DATA_BLOCK "DB_SDC_TS_PARAMETER_6"   // DB3709
{ S7_Optimized_Access := 'FALSE' }
AUTHOR : FFM
FAMILY : SDC
NAME : SECT_DEF
VERSION : 1.0
   VAR
      HEADER : Struct   // Struktur für Datenheader // nicht verschieben
         DB_NR : Int := 3709;   // DB Nummer
         MIN_NR_SEK : Int := 501;   // Niedrigste SEK Nummer im DB
         MAX_NR_SEK : Int := 600;   // Höchste SEK Nummer im DB
         START_DAT : Int := 20;   // Startadresse der SEK im DB
         LAENGE_SEK_DATA : Int := 260;   // Länge SEK Data
         ANZ_PROFIL : Int := 10;   // Number of Profiles
         OFFEST_PROFIL : Int := 40;   // Offestadresse der Profilparameter im TS-Parameterdatensatz
         LAENGE_PROFIL_DATA : Int := 22;   // Länge SEK Data
         Res160 : Int := 0;   // Reserve
         Res : Int := 0;   // Reserve
      END_STRUCT;
      TS : Array[501..600] of "UDT_SDC_TS_PARAMETER";
   END_VAR
BEGIN
   TS[501].ALLG.SEK_NEXT_1 := 0;
   TS[501].ALLG.SEK_NEXT_2 := 0;
   TS[501].ALLG.Spare[4] := 16#00;
   TS[501].ALLG.Spare[5] := 16#00;
   TS[501].ALLG.POS.Start_1 := 1639750;
   TS[501].ALLG.POS.End_1 := 1646749;
   TS[501].ALLG.POS.Start_2 := 0;
   TS[501].ALLG.POS.End_2 := 0;
   TS[501].ALLG.POS.Actionpoint_1 := 0;
   TS[501].ALLG.POS.Actionpoint_2 := 0;
   TS[501].ALLG.FLAGS.DIST_VAL[0] := FALSE;
   TS[501].ALLG.FLAGS.DIST_VAL[1] := FALSE;
   TS[501].ALLG.FLAGS.DIST_VAL[2] := FALSE;
   TS[501].ALLG.FLAGS.DIST_VAL[3] := FALSE;
   TS[501].ALLG.FLAGS.DIST_VAL[4] := FALSE;
   TS[501].ALLG.FLAGS.DIST_VAL[5] := FALSE;
   TS[501].ALLG.FLAGS.DIST_VAL[6] := FALSE;
   TS[501].ALLG.FLAGS.DIST_VAL[7] := FALSE;
   TS[501].ALLG.FLAGS.DIST_VAL[8] := FALSE;
   TS[501].ALLG.FLAGS.DIST_VAL[9] := TRUE;
   TS[501].ALLG.FLAGS.DIST_VAL[10] := FALSE;
   TS[501].ALLG.FLAGS.DIST_VAL[11] := FALSE;
   TS[501].ALLG.FLAGS.DIST_VAL[12] := FALSE;
   TS[501].ALLG.FLAGS.DIST_VAL[13] := FALSE;
   TS[501].ALLG.FLAGS.DIST_VAL[14] := FALSE;
   TS[501].ALLG.FLAGS.DIST_VAL[15] := FALSE;
   TS[501].ALLG.FLAGS.one_profile := FALSE;
   TS[501].ALLG.FLAGS.BLIND := FALSE;
   TS[501].ALLG.FLAGS.NO_DIST_CONT := FALSE;
   TS[501].ALLG.FLAGS.SYNCH_AREA := FALSE;
   TS[501].ALLG.FLAGS.bit24 := FALSE;
   TS[501].ALLG.FLAGS.bit25 := FALSE;
   TS[501].ALLG.FLAGS.bit26 := FALSE;
   TS[501].ALLG.FLAGS.bit27 := FALSE;
   TS[501].ALLG.FLAGS.EN_HOIST := FALSE;
   TS[501].ALLG.FLAGS.D_RESET_AFTER := FALSE;
   TS[501].ALLG.FLAGS.D_PULK := FALSE;
   TS[501].ALLG.FLAGS.bit33 := FALSE;
   TS[501].ALLG.FLAGS.bit34 := FALSE;
   TS[501].ALLG.FLAGS.bit35 := FALSE;
   TS[501].ALLG.FLAGS.bit36 := FALSE;
   TS[501].ALLG.FLAGS.Deutronic_ON := FALSE;
   TS[501].ALLG.Stop_Position := 6500;
   TS[501].ALLG.Drive_speed_1 := 15000;
   TS[501].ALLG.Drive_speed_2 := 6000;
   TS[501].PROFIL[1].Hoist_Pos_start := 0;
   TS[501].PROFIL[1].Height := 3890;
   TS[501].PROFIL[1].Hoist_speed := 2000;
   TS[501].PROFIL[1].Hoist_offset_1 := 0;
   TS[501].PROFIL[1].Hoist_offset_2 := 0;
   TS[501].PROFIL[1].Hoist_offset_3 := 0;
   TS[501].PROFIL[1].Hoist_offset_4 := 0;
   TS[501].PROFIL[1].Hoist_Start_offset_1 := 0;
   TS[501].PROFIL[1].Hoist_Start_offset_2 := 0;
   TS[501].PROFIL[1].Hoist_Start_offset_3 := 0;
   TS[501].PROFIL[1].Hoist_Start_offset_4 := 0;
   TS[501].PROFIL[2].Hoist_Pos_start := 0;
   TS[501].PROFIL[2].Height := 3890;
   TS[501].PROFIL[2].Hoist_speed := 2000;
   TS[501].PROFIL[2].Hoist_offset_1 := 0;
   TS[501].PROFIL[2].Hoist_offset_2 := 0;
   TS[501].PROFIL[2].Hoist_offset_3 := 0;
   TS[501].PROFIL[2].Hoist_offset_4 := 0;
   TS[501].PROFIL[2].Hoist_Start_offset_1 := 0;
   TS[501].PROFIL[2].Hoist_Start_offset_2 := 0;
   TS[501].PROFIL[2].Hoist_Start_offset_3 := 0;
   TS[501].PROFIL[2].Hoist_Start_offset_4 := 0;
   TS[501].PROFIL[3].Hoist_Pos_start := 0;
   TS[501].PROFIL[3].Height := 3890;
   TS[501].PROFIL[3].Hoist_speed := 2000;
   TS[501].PROFIL[3].Hoist_offset_1 := 0;
   TS[501].PROFIL[3].Hoist_offset_2 := 0;
   TS[501].PROFIL[3].Hoist_offset_3 := 0;
   TS[501].PROFIL[3].Hoist_offset_4 := 0;
   TS[501].PROFIL[3].Hoist_Start_offset_1 := 0;
   TS[501].PROFIL[3].Hoist_Start_offset_2 := 0;
   TS[501].PROFIL[3].Hoist_Start_offset_3 := 0;
   TS[501].PROFIL[3].Hoist_Start_offset_4 := 0;
   TS[501].PROFIL[4].Hoist_Pos_start := 0;
   TS[501].PROFIL[4].Height := 3890;
   TS[501].PROFIL[4].Hoist_speed := 2000;
   TS[501].PROFIL[4].Hoist_offset_1 := 0;
   TS[501].PROFIL[4].Hoist_offset_2 := 0;
   TS[501].PROFIL[4].Hoist_offset_3 := 0;
   TS[501].PROFIL[4].Hoist_offset_4 := 0;
   TS[501].PROFIL[4].Hoist_Start_offset_1 := 0;
   TS[501].PROFIL[4].Hoist_Start_offset_2 := 0;
   TS[501].PROFIL[4].Hoist_Start_offset_3 := 0;
   TS[501].PROFIL[4].Hoist_Start_offset_4 := 0;
   TS[501].PROFIL[5].Hoist_Pos_start := 0;
   TS[501].PROFIL[5].Height := 3890;
   TS[501].PROFIL[5].Hoist_speed := 2000;
   TS[501].PROFIL[5].Hoist_offset_1 := 0;
   TS[501].PROFIL[5].Hoist_offset_2 := 0;
   TS[501].PROFIL[5].Hoist_offset_3 := 0;
   TS[501].PROFIL[5].Hoist_offset_4 := 0;
   TS[501].PROFIL[5].Hoist_Start_offset_1 := 0;
   TS[501].PROFIL[5].Hoist_Start_offset_2 := 0;
   TS[501].PROFIL[5].Hoist_Start_offset_3 := 0;
   TS[501].PROFIL[5].Hoist_Start_offset_4 := 0;
   TS[501].PROFIL[6].Hoist_Pos_start := 0;
   TS[501].PROFIL[6].Height := 3890;
   TS[501].PROFIL[6].Hoist_speed := 2000;
   TS[501].PROFIL[6].Hoist_offset_1 := 0;
   TS[501].PROFIL[6].Hoist_offset_2 := 0;
   TS[501].PROFIL[6].Hoist_offset_3 := 0;
   TS[501].PROFIL[6].Hoist_offset_4 := 0;
   TS[501].PROFIL[6].Hoist_Start_offset_1 := 0;
   TS[501].PROFIL[6].Hoist_Start_offset_2 := 0;
   TS[501].PROFIL[6].Hoist_Start_offset_3 := 0;
   TS[501].PROFIL[6].Hoist_Start_offset_4 := 0;
   TS[501].PROFIL[7].Hoist_Pos_start := 0;
   TS[501].PROFIL[7].Height := 3890;
   TS[501].PROFIL[7].Hoist_speed := 2000;
   TS[501].PROFIL[7].Hoist_offset_1 := 0;
   TS[501].PROFIL[7].Hoist_offset_2 := 0;
   TS[501].PROFIL[7].Hoist_offset_3 := 0;
   TS[501].PROFIL[7].Hoist_offset_4 := 0;
   TS[501].PROFIL[7].Hoist_Start_offset_1 := 0;
   TS[501].PROFIL[7].Hoist_Start_offset_2 := 0;
   TS[501].PROFIL[7].Hoist_Start_offset_3 := 0;
   TS[501].PROFIL[7].Hoist_Start_offset_4 := 0;
   TS[501].PROFIL[8].Hoist_Pos_start := 0;
   TS[501].PROFIL[8].Height := 3890;
   TS[501].PROFIL[8].Hoist_speed := 2000;
   TS[501].PROFIL[8].Hoist_offset_1 := 0;
   TS[501].PROFIL[8].Hoist_offset_2 := 0;
   TS[501].PROFIL[8].Hoist_offset_3 := 0;
   TS[501].PROFIL[8].Hoist_offset_4 := 0;
   TS[501].PROFIL[8].Hoist_Start_offset_1 := 0;
   TS[501].PROFIL[8].Hoist_Start_offset_2 := 0;
   TS[501].PROFIL[8].Hoist_Start_offset_3 := 0;
   TS[501].PROFIL[8].Hoist_Start_offset_4 := 0;
   TS[501].PROFIL[9].Hoist_Pos_start := 0;
   TS[501].PROFIL[9].Height := 3890;
   TS[501].PROFIL[9].Hoist_speed := 2000;
   TS[501].PROFIL[9].Hoist_offset_1 := 0;
   TS[501].PROFIL[9].Hoist_offset_2 := 0;
   TS[501].PROFIL[9].Hoist_offset_3 := 0;
   TS[501].PROFIL[9].Hoist_offset_4 := 0;
   TS[501].PROFIL[9].Hoist_Start_offset_1 := 0;
   TS[501].PROFIL[9].Hoist_Start_offset_2 := 0;
   TS[501].PROFIL[9].Hoist_Start_offset_3 := 0;
   TS[501].PROFIL[9].Hoist_Start_offset_4 := 0;
   TS[501].PROFIL[10].Hoist_Pos_start := 0;
   TS[501].PROFIL[10].Height := 3890;
   TS[501].PROFIL[10].Hoist_speed := 2000;
   TS[501].PROFIL[10].Hoist_offset_1 := 0;
   TS[501].PROFIL[10].Hoist_offset_2 := 0;
   TS[501].PROFIL[10].Hoist_offset_3 := 0;
   TS[501].PROFIL[10].Hoist_offset_4 := 0;
   TS[501].PROFIL[10].Hoist_Start_offset_1 := 0;
   TS[501].PROFIL[10].Hoist_Start_offset_2 := 0;
   TS[501].PROFIL[10].Hoist_Start_offset_3 := 0;
   TS[501].PROFIL[10].Hoist_Start_offset_4 := 0;
   TS[502].ALLG.SEK_NEXT_1 := 0;
   TS[502].ALLG.SEK_NEXT_2 := 0;
   TS[502].ALLG.Spare[4] := 16#00;
   TS[502].ALLG.Spare[5] := 16#00;
   TS[502].ALLG.POS.Start_1 := 1646750;
   TS[502].ALLG.POS.End_1 := 1653749;
   TS[502].ALLG.POS.Start_2 := 0;
   TS[502].ALLG.POS.End_2 := 0;
   TS[502].ALLG.POS.Actionpoint_1 := 0;
   TS[502].ALLG.POS.Actionpoint_2 := 0;
   TS[502].ALLG.FLAGS.DIST_VAL[0] := FALSE;
   TS[502].ALLG.FLAGS.DIST_VAL[1] := FALSE;
   TS[502].ALLG.FLAGS.DIST_VAL[2] := FALSE;
   TS[502].ALLG.FLAGS.DIST_VAL[3] := FALSE;
   TS[502].ALLG.FLAGS.DIST_VAL[4] := FALSE;
   TS[502].ALLG.FLAGS.DIST_VAL[5] := FALSE;
   TS[502].ALLG.FLAGS.DIST_VAL[6] := FALSE;
   TS[502].ALLG.FLAGS.DIST_VAL[7] := FALSE;
   TS[502].ALLG.FLAGS.DIST_VAL[8] := FALSE;
   TS[502].ALLG.FLAGS.DIST_VAL[9] := TRUE;
   TS[502].ALLG.FLAGS.DIST_VAL[10] := FALSE;
   TS[502].ALLG.FLAGS.DIST_VAL[11] := FALSE;
   TS[502].ALLG.FLAGS.DIST_VAL[12] := FALSE;
   TS[502].ALLG.FLAGS.DIST_VAL[13] := FALSE;
   TS[502].ALLG.FLAGS.DIST_VAL[14] := FALSE;
   TS[502].ALLG.FLAGS.DIST_VAL[15] := FALSE;
   TS[502].ALLG.FLAGS.one_profile := FALSE;
   TS[502].ALLG.FLAGS.BLIND := FALSE;
   TS[502].ALLG.FLAGS.NO_DIST_CONT := FALSE;
   TS[502].ALLG.FLAGS.SYNCH_AREA := FALSE;
   TS[502].ALLG.FLAGS.bit24 := FALSE;
   TS[502].ALLG.FLAGS.bit25 := FALSE;
   TS[502].ALLG.FLAGS.bit26 := FALSE;
   TS[502].ALLG.FLAGS.bit27 := FALSE;
   TS[502].ALLG.FLAGS.EN_HOIST := FALSE;
   TS[502].ALLG.FLAGS.D_RESET_AFTER := FALSE;
   TS[502].ALLG.FLAGS.D_PULK := FALSE;
   TS[502].ALLG.FLAGS.bit33 := FALSE;
   TS[502].ALLG.FLAGS.bit34 := FALSE;
   TS[502].ALLG.FLAGS.bit35 := FALSE;
   TS[502].ALLG.FLAGS.bit36 := FALSE;
   TS[502].ALLG.FLAGS.Deutronic_ON := FALSE;
   TS[502].ALLG.Stop_Position := 6400;
   TS[502].ALLG.Drive_speed_1 := 15000;
   TS[502].ALLG.Drive_speed_2 := 6000;
   // 15300 more start values not shown
END_DATA_BLOCK

DATA_BLOCK "DB_SDC_EMS_1"   // DB3714
{ S7_Optimized_Access := 'FALSE' }
VERSION : 0.1
   VAR
      HEADER : Struct
         DB_NR : Int := 3714;
         MIN_NR_EMS : Int := 1;
         MAX_NR_EMS : Int := 200;
         START_EMS : Int := 20;
         LAENGE_EMS : Int := 260;
         OFFSET_EMS_SEK_STAT : Int := 164;
         LAENGE_EMS_SEK_STAT : Int := 34;
         OFFSET_EMS_FKT : Int := 216;
         Res160 : Int := 0;
         Load : Bool := TRUE;
      END_STRUCT;
   END_VAR
BEGIN
END_DATA_BLOCK

DATA_BLOCK "DB_SDC_TS_IF_COMMAND"   // DB3716
{ S7_Optimized_Access := 'FALSE' }
AUTHOR : FFM
FAMILY : SDC
NAME : SECT_IF
VERSION : 0.1
   VAR
      HEADER : Struct   // Struktur für Datenheader // nicht verschieben
         DB_NR : Int := 3716;   // DB Nummer
         MIN_NR_SEK : Int := 1;   // Niedrigste SEK Nummer im DB
         MAX_NR_SEK : Int := 600;   // Höchste SEK Nummer im DB
         START_DAT : Int := 20;   // Startadresse der SEK im DB
         LAENGE_SEK_DATA : Int := 18;   // Länge SEK Data
         LAENGE_VAL_DATA : Int := 8;   // Länge Value Data
         LAENGE_BIT_DATA : Int := 6;   // Länge Bit Data
         LAENGE_FKT : Int := 4;   // Länge Funktion
         Res16 : Int;   // Reserve
         Res18 : Int;   // Reserve
      END_STRUCT;
      SEK : Array[1..600] of "UDT_SDC_EMS_TS_COM";   // Komando für Sektion
   END_VAR
BEGIN
END_DATA_BLOCK

DATA_BLOCK "DB_SDC_TS_IF_COMMAND_2"   // DB3717
{ S7_Optimized_Access := 'FALSE' }
AUTHOR : FFM
FAMILY : SDC
NAME : SECT_IF
VERSION : 0.1
   VAR
      HEADER : Struct   // Struktur für Datenheader // nicht verschieben
         DB_NR : Int := 3717;   // DB Nummer
         MIN_NR_SEK : Int := 601;   // Niedrigste SEK Nummer im DB
         MAX_NR_SEK : Int := 1000;   // Höchste SEK Nummer im DB
         START_DAT : Int := 20;   // Startadresse der SEK im DB
         LAENGE_SEK_DATA : Int := 18;   // Länge SEK Data
         LAENGE_VAL_DATA : Int := 8;   // Länge Value Data
         LAENGE_BIT_DATA : Int := 6;   // Länge Bit Data
         LAENGE_FKT : Int := 4;   // Länge Funktion
         Res16 : Int;   // Reserve
         Res18 : Int;   // Reserve
      END_STRUCT;
      SEK : Array[601..1000] of "UDT_SDC_EMS_TS_COM";   // Komando für Sektion
   END_VAR
BEGIN
END_DATA_BLOCK

DATA_BLOCK "DB_SDC_TS_IF_STATUS"   // DB3718
{ S7_Optimized_Access := 'FALSE' }
AUTHOR : FFM
FAMILY : SDC
NAME : SECT_IF
VERSION : 1.0
   VAR
      HEADER : Struct
         DB_NR : Int := 3718;
         MIN_NR_SEK : Int := 1;
         MAX_NR_SEK : Int := 600;
         START_DAT : Int := 20;
         LAENGE_SEK_DATA : Int := 34;
         LAENGE_VAL_DATA : Int := 18;
         LAENGE_BIT_DATA : Int := 8;
         LAENGE_SERIES : Int := 4;
         LAENGE_FKT : Int := 4;
         Res18 : Int := 0;
      END_STRUCT;
      SEK : Array[1..600] of "UDT_SDC_EMS_TS_STAT";
   END_VAR
BEGIN
   SEK[1].VAL.EMS_ID := 1;
   SEK[1].VAL.PROFIL := 1;
   SEK[1].VAL.DRIVE_POS := 581346;
   SEK[1].VAL.HOIST_POS := 4151;
   SEK[1].VAL.ERROR := 504;
   SEK[1].VAL.DRIVE_POS_PERC := 0;
   SEK[1].VAL.SEK := 1;
   SEK[1].BIT.PRESENT := TRUE;
   SEK[1].BIT.ERROR := TRUE;
   SEK[1].BIT.MAN_IR := TRUE;
   SEK[1].BIT.MORE_EMS_PRESENT := FALSE;
   SEK[1].BIT.ER_COMMAND := FALSE;
   SEK[1].BIT.W_DIST := FALSE;
   SEK[1].BIT.Spare_0_6 := FALSE;
   SEK[1].BIT.MESS_ACT := FALSE;
   SEK[1].BIT.D_MOVING := FALSE;
   SEK[1].BIT.D_NOT_MOVING := TRUE;
   SEK[1].BIT.H_MOVING := FALSE;
   SEK[1].BIT.H_NOT_MOVING := TRUE;
   SEK[1].BIT.X_MOVING := FALSE;
   SEK[1].BIT.X_NOT_MOVING := TRUE;
   SEK[1].BIT.D_IN_POS := FALSE;
   SEK[1].BIT.Spare_2_1 := FALSE;
   SEK[1].BIT.D_BEFOR_POS := FALSE;
   SEK[1].BIT.D_AFTER_POS := TRUE;
   SEK[1].BIT.D_GR_AP1 := TRUE;
   SEK[1].BIT.D_SM_AP1 := FALSE;
   SEK[1].BIT.D_GR_AP2 := TRUE;
   SEK[1].BIT.D_SM_AP2 := FALSE;
   SEK[1].BIT.H_IN_POS := TRUE;
   SEK[1].BIT.H_IN_TOPPOS := TRUE;
   SEK[1].BIT.H_IN_POS1 := FALSE;
   SEK[1].BIT.H_IN_POS2 := FALSE;
   SEK[1].BIT.H_IN_POS3 := FALSE;
   SEK[1].BIT.H_IN_POS4 := FALSE;
   SEK[1].BIT.H_GR_POS := FALSE;
   SEK[1].BIT.H_SM_POS := FALSE;
   SEK[1].BIT.H_GR_POS1 := FALSE;
   SEK[1].BIT.H_SM_POS1 := FALSE;
   SEK[1].BIT.H_GR_POS2 := FALSE;
   SEK[1].BIT.H_SM_POS2 := FALSE;
   SEK[1].BIT.H_GR_POS3 := FALSE;
   SEK[1].BIT.H_SM_POS3 := FALSE;
   SEK[1].BIT.H_GR_POS4 := FALSE;
   SEK[1].BIT.H_SM_POS4 := FALSE;
   SEK[1].BIT.H_BOTTOM_POS := FALSE;
   SEK[1].BIT.H_DISABLED := TRUE;
   SEK[1].BIT.H_CLEAR := FALSE;
   SEK[1].BIT.D_MOVING_FWD := FALSE;
   SEK[1].BIT.D_MOVING_RWD := FALSE;
   SEK[1].BIT.D_RESET_AFTER := FALSE;
   SEK[1].BIT.D_PULK := FALSE;
   SEK[1].BIT.D_NO_POS := FALSE;
   SEK[1].SORTE[1] := 'L';
   SEK[1].SORTE[2] := 'E';
   SEK[1].SORTE[3] := 'E';
   SEK[1].SORTE[4] := 'R';
   SEK[1].FKT.EMS_TO_REPAIR_1 := FALSE;
   SEK[1].FKT.EMS_TO_REPAIR_2 := FALSE;
   SEK[1].FKT.EMERG_HOIST := FALSE;
   SEK[1].FKT.Reserve_03 := FALSE;
   SEK[1].FKT.EMERG_DRIVE_FC := FALSE;
   SEK[1].FKT.Reserve_05 := FALSE;
   SEK[1].FKT.LAMP_TEST := FALSE;
   SEK[1].FKT.VAC_CLEAN := FALSE;
   SEK[1].FKT.PE_TEST := FALSE;
   SEK[1].FKT.KOHLE_TEST := FALSE;
   SEK[1].FKT.KOM_TEST := FALSE;
   SEK[1].FKT.Reserve_11 := FALSE;
   SEK[1].FKT.Reserve_12 := FALSE;
   SEK[1].FKT.Reserve_13 := FALSE;
   SEK[1].FKT.Reserve_14 := FALSE;
   SEK[1].FKT.Reserve_15 := FALSE;
   SEK[1].SPARE := 16#0000;
   SEK[2].VAL.EMS_ID := 0;
   SEK[2].VAL.PROFIL := 0;
   SEK[2].VAL.DRIVE_POS := 0;
   SEK[2].VAL.HOIST_POS := 0;
   SEK[2].VAL.ERROR := 0;
   SEK[2].VAL.DRIVE_POS_PERC := 0;
   SEK[2].VAL.SEK := 0;
   SEK[2].BIT.PRESENT := FALSE;
   SEK[2].BIT.ERROR := FALSE;
   SEK[2].BIT.MAN_IR := FALSE;
   SEK[2].BIT.MORE_EMS_PRESENT := FALSE;
   SEK[2].BIT.ER_COMMAND := FALSE;
   SEK[2].BIT.W_DIST := FALSE;
   SEK[2].BIT.Spare_0_6 := FALSE;
   SEK[2].BIT.MESS_ACT := FALSE;
   SEK[2].BIT.D_MOVING := FALSE;
   SEK[2].BIT.D_NOT_MOVING := FALSE;
   SEK[2].BIT.H_MOVING := FALSE;
   SEK[2].BIT.H_NOT_MOVING := FALSE;
   SEK[2].BIT.X_MOVING := FALSE;
   SEK[2].BIT.X_NOT_MOVING := FALSE;
   SEK[2].BIT.D_IN_POS := FALSE;
   SEK[2].BIT.Spare_2_1 := FALSE;
   SEK[2].BIT.D_BEFOR_POS := FALSE;
   SEK[2].BIT.D_AFTER_POS := FALSE;
   SEK[2].BIT.D_GR_AP1 := FALSE;
   SEK[2].BIT.D_SM_AP1 := FALSE;
   SEK[2].BIT.D_GR_AP2 := FALSE;
   SEK[2].BIT.D_SM_AP2 := FALSE;
   SEK[2].BIT.H_IN_POS := FALSE;
   SEK[2].BIT.H_IN_TOPPOS := FALSE;
   SEK[2].BIT.H_IN_POS1 := FALSE;
   SEK[2].BIT.H_IN_POS2 := FALSE;
   SEK[2].BIT.H_IN_POS3 := FALSE;
   SEK[2].BIT.H_IN_POS4 := FALSE;
   SEK[2].BIT.H_GR_POS := FALSE;
   SEK[2].BIT.H_SM_POS := FALSE;
   SEK[2].BIT.H_GR_POS1 := FALSE;
   SEK[2].BIT.H_SM_POS1 := FALSE;
   SEK[2].BIT.H_GR_POS2 := FALSE;
   SEK[2].BIT.H_SM_POS2 := FALSE;
   SEK[2].BIT.H_GR_POS3 := FALSE;
   SEK[2].BIT.H_SM_POS3 := FALSE;
   SEK[2].BIT.H_GR_POS4 := FALSE;
   SEK[2].BIT.H_SM_POS4 := FALSE;
   SEK[2].BIT.H_BOTTOM_POS := FALSE;
   SEK[2].BIT.H_DISABLED := FALSE;
   SEK[2].BIT.H_CLEAR := FALSE;
   SEK[2].BIT.D_MOVING_FWD := FALSE;
   SEK[2].BIT.D_MOVING_RWD := FALSE;
   SEK[2].BIT.D_RESET_AFTER := FALSE;
   SEK[2].BIT.D_PULK := FALSE;
   SEK[2].BIT.D_NO_POS := TRUE;
   SEK[2].SORTE[1] := ' ';
   SEK[2].SORTE[2] := ' ';
   SEK[2].SORTE[3] := ' ';
   SEK[2].SORTE[4] := ' ';
   SEK[2].FKT.EMS_TO_REPAIR_1 := FALSE;
   SEK[2].FKT.EMS_TO_REPAIR_2 := FALSE;
   SEK[2].FKT.EMERG_HOIST := FALSE;
   SEK[2].FKT.Reserve_03 := FALSE;
   SEK[2].FKT.EMERG_DRIVE_FC := FALSE;
   SEK[2].FKT.Reserve_05 := FALSE;
   SEK[2].FKT.LAMP_TEST := FALSE;
   SEK[2].FKT.VAC_CLEAN := FALSE;
   SEK[2].FKT.PE_TEST := FALSE;
   SEK[2].FKT.KOHLE_TEST := FALSE;
   SEK[2].FKT.KOM_TEST := FALSE;
   SEK[2].FKT.Reserve_11 := FALSE;
   SEK[2].FKT.Reserve_12 := FALSE;
   SEK[2].FKT.Reserve_13 := FALSE;
   SEK[2].FKT.Reserve_14 := FALSE;
   SEK[2].FKT.Reserve_15 := FALSE;
   SEK[2].SPARE := 16#0000;
   SEK[3].VAL.EMS_ID := 0;
   SEK[3].VAL.PROFIL := 0;
   SEK[3].VAL.DRIVE_POS := 0;
   SEK[3].VAL.HOIST_POS := 0;
   SEK[3].VAL.ERROR := 0;
   SEK[3].VAL.DRIVE_POS_PERC := 0;
   SEK[3].VAL.SEK := 0;
   SEK[3].BIT.PRESENT := FALSE;
   SEK[3].BIT.ERROR := FALSE;
   SEK[3].BIT.MAN_IR := FALSE;
   SEK[3].BIT.MORE_EMS_PRESENT := FALSE;
   SEK[3].BIT.ER_COMMAND := FALSE;
   SEK[3].BIT.W_DIST := FALSE;
   SEK[3].BIT.Spare_0_6 := FALSE;
   SEK[3].BIT.MESS_ACT := FALSE;
   SEK[3].BIT.D_MOVING := FALSE;
   SEK[3].BIT.D_NOT_MOVING := FALSE;
   SEK[3].BIT.H_MOVING := FALSE;
   SEK[3].BIT.H_NOT_MOVING := FALSE;
   SEK[3].BIT.X_MOVING := FALSE;
   SEK[3].BIT.X_NOT_MOVING := FALSE;
   SEK[3].BIT.D_IN_POS := FALSE;
   SEK[3].BIT.Spare_2_1 := FALSE;
   SEK[3].BIT.D_BEFOR_POS := FALSE;
   SEK[3].BIT.D_AFTER_POS := FALSE;
   SEK[3].BIT.D_GR_AP1 := FALSE;
   SEK[3].BIT.D_SM_AP1 := FALSE;
   SEK[3].BIT.D_GR_AP2 := FALSE;
   SEK[3].BIT.D_SM_AP2 := FALSE;
   SEK[3].BIT.H_IN_POS := FALSE;
   SEK[3].BIT.H_IN_TOPPOS := FALSE;
   SEK[3].BIT.H_IN_POS1 := FALSE;
   SEK[3].BIT.H_IN_POS2 := FALSE;
   SEK[3].BIT.H_IN_POS3 := FALSE;
   SEK[3].BIT.H_IN_POS4 := FALSE;
   SEK[3].BIT.H_GR_POS := FALSE;
   SEK[3].BIT.H_SM_POS := FALSE;
   SEK[3].BIT.H_GR_POS1 := FALSE;
   SEK[3].BIT.H_SM_POS1 := FALSE;
   SEK[3].BIT.H_GR_POS2 := FALSE;
   SEK[3].BIT.H_SM_POS2 := FALSE;
   SEK[3].BIT.H_GR_POS3 := FALSE;
   SEK[3].BIT.H_SM_POS3 := FALSE;
   SEK[3].BIT.H_GR_POS4 := FALSE;
   SEK[3].BIT.H_SM_POS4 := FALSE;
   SEK[3].BIT.H_BOTTOM_POS := FALSE;
   SEK[3].BIT.H_DISABLED := FALSE;
   SEK[3].BIT.H_CLEAR := FALSE;
   SEK[3].BIT.D_MOVING_FWD := FALSE;
   SEK[3].BIT.D_MOVING_RWD := FALSE;
   SEK[3].BIT.D_RESET_AFTER := FALSE;
   SEK[3].BIT.D_PULK := FALSE;
   // 44200 more start values not shown
END_DATA_BLOCK

DATA_BLOCK "DB_SDC_TS_IF_STATUS_2"   // DB3719
{ S7_Optimized_Access := 'FALSE' }
AUTHOR : FFM
FAMILY : SDC
NAME : SECT_IF
VERSION : 1.0
   VAR
      HEADER : Struct   // Struktur für Datenheader // nicht verschieben
         DB_NR : Int := 3719;   // DB Nummer
         MIN_NR_SEK : Int := 601;   // Niedrigste SEK Nummer im DB
         MAX_NR_SEK : Int := 1000;   // Höchste SEK Nummer im DB
         START_DAT : Int := 20;   // Startadresse der SEK im DB
         LAENGE_SEK_DATA : Int := 34;   // Länge SEK Data
         LAENGE_VAL_DATA : Int := 18;   // Länge Value Data
         LAENGE_BIT_DATA : Int := 8;   // Länge Bit Data
         LAENGE_SERIES : Int := 4;   // Länge SERIES
         LAENGE_FKT : Int := 4;   // Länge Funktion
         Res18 : Int := 0;   // Reserve
      END_STRUCT;
      SEK : Array[601..1000] of "UDT_SDC_EMS_TS_STAT";   // Status of section
   END_VAR
BEGIN
   SEK[601].VAL.EMS_ID := 0;
   SEK[601].VAL.PROFIL := 0;
   SEK[601].VAL.DRIVE_POS := 0;
   SEK[601].VAL.HOIST_POS := 0;
   SEK[601].VAL.ERROR := 0;
   SEK[601].VAL.DRIVE_POS_PERC := 0;
   SEK[601].VAL.SEK := 0;
   SEK[601].BIT.PRESENT := FALSE;
   SEK[601].BIT.ERROR := FALSE;
   SEK[601].BIT.MAN_IR := FALSE;
   SEK[601].BIT.MORE_EMS_PRESENT := FALSE;
   SEK[601].BIT.ER_COMMAND := FALSE;
   SEK[601].BIT.W_DIST := FALSE;
   SEK[601].BIT.Spare_0_6 := FALSE;
   SEK[601].BIT.MESS_ACT := FALSE;
   SEK[601].BIT.D_MOVING := FALSE;
   SEK[601].BIT.D_NOT_MOVING := FALSE;
   SEK[601].BIT.H_MOVING := FALSE;
   SEK[601].BIT.H_NOT_MOVING := FALSE;
   SEK[601].BIT.X_MOVING := FALSE;
   SEK[601].BIT.X_NOT_MOVING := FALSE;
   SEK[601].BIT.D_IN_POS := FALSE;
   SEK[601].BIT.Spare_2_1 := FALSE;
   SEK[601].BIT.D_BEFOR_POS := FALSE;
   SEK[601].BIT.D_AFTER_POS := FALSE;
   SEK[601].BIT.D_GR_AP1 := FALSE;
   SEK[601].BIT.D_SM_AP1 := FALSE;
   SEK[601].BIT.D_GR_AP2 := FALSE;
   SEK[601].BIT.D_SM_AP2 := FALSE;
   SEK[601].BIT.H_IN_POS := FALSE;
   SEK[601].BIT.H_IN_TOPPOS := FALSE;
   SEK[601].BIT.H_IN_POS1 := FALSE;
   SEK[601].BIT.H_IN_POS2 := FALSE;
   SEK[601].BIT.H_IN_POS3 := FALSE;
   SEK[601].BIT.H_IN_POS4 := FALSE;
   SEK[601].BIT.H_GR_POS := FALSE;
   SEK[601].BIT.H_SM_POS := FALSE;
   SEK[601].BIT.H_GR_POS1 := FALSE;
   SEK[601].BIT.H_SM_POS1 := FALSE;
   SEK[601].BIT.H_GR_POS2 := FALSE;
   SEK[601].BIT.H_SM_POS2 := FALSE;
   SEK[601].BIT.H_GR_POS3 := FALSE;
   SEK[601].BIT.H_SM_POS3 := FALSE;
   SEK[601].BIT.H_GR_POS4 := FALSE;
   SEK[601].BIT.H_SM_POS4 := FALSE;
   SEK[601].BIT.H_BOTTOM_POS := FALSE;
   SEK[601].BIT.H_DISABLED := FALSE;
   SEK[601].BIT.H_CLEAR := FALSE;
   SEK[601].BIT.D_MOVING_FWD := FALSE;
   SEK[601].BIT.D_MOVING_RWD := FALSE;
   SEK[601].BIT.D_RESET_AFTER := FALSE;
   SEK[601].BIT.D_PULK := FALSE;
   SEK[601].BIT.D_NO_POS := FALSE;
   SEK[601].SORTE[1] := ' ';
   SEK[601].SORTE[2] := ' ';
   SEK[601].SORTE[3] := ' ';
   SEK[601].SORTE[4] := ' ';
   SEK[601].FKT.EMS_TO_REPAIR_1 := FALSE;
   SEK[601].FKT.EMS_TO_REPAIR_2 := FALSE;
   SEK[601].FKT.EMERG_HOIST := FALSE;
   SEK[601].FKT.Reserve_03 := FALSE;
   SEK[601].FKT.EMERG_DRIVE_FC := FALSE;
   SEK[601].FKT.Reserve_05 := FALSE;
   SEK[601].FKT.LAMP_TEST := FALSE;
   SEK[601].FKT.VAC_CLEAN := FALSE;
   SEK[601].FKT.PE_TEST := FALSE;
   SEK[601].FKT.KOHLE_TEST := FALSE;
   SEK[601].FKT.KOM_TEST := FALSE;
   SEK[601].FKT.Reserve_11 := FALSE;
   SEK[601].FKT.Reserve_12 := FALSE;
   SEK[601].FKT.Reserve_13 := FALSE;
   SEK[601].FKT.Reserve_14 := FALSE;
   SEK[601].FKT.Reserve_15 := FALSE;
   SEK[601].SPARE := 16#0000;
   SEK[602].VAL.EMS_ID := 0;
   SEK[602].VAL.PROFIL := 0;
   SEK[602].VAL.DRIVE_POS := 0;
   SEK[602].VAL.HOIST_POS := 0;
   SEK[602].VAL.ERROR := 0;
   SEK[602].VAL.DRIVE_POS_PERC := 0;
   SEK[602].VAL.SEK := 0;
   SEK[602].BIT.PRESENT := FALSE;
   SEK[602].BIT.ERROR := FALSE;
   SEK[602].BIT.MAN_IR := FALSE;
   SEK[602].BIT.MORE_EMS_PRESENT := FALSE;
   SEK[602].BIT.ER_COMMAND := FALSE;
   SEK[602].BIT.W_DIST := FALSE;
   SEK[602].BIT.Spare_0_6 := FALSE;
   SEK[602].BIT.MESS_ACT := FALSE;
   SEK[602].BIT.D_MOVING := FALSE;
   SEK[602].BIT.D_NOT_MOVING := FALSE;
   SEK[602].BIT.H_MOVING := FALSE;
   SEK[602].BIT.H_NOT_MOVING := FALSE;
   SEK[602].BIT.X_MOVING := FALSE;
   SEK[602].BIT.X_NOT_MOVING := FALSE;
   SEK[602].BIT.D_IN_POS := FALSE;
   SEK[602].BIT.Spare_2_1 := FALSE;
   SEK[602].BIT.D_BEFOR_POS := FALSE;
   SEK[602].BIT.D_AFTER_POS := FALSE;
   SEK[602].BIT.D_GR_AP1 := FALSE;
   SEK[602].BIT.D_SM_AP1 := FALSE;
   SEK[602].BIT.D_GR_AP2 := FALSE;
   SEK[602].BIT.D_SM_AP2 := FALSE;
   SEK[602].BIT.H_IN_POS := FALSE;
   SEK[602].BIT.H_IN_TOPPOS := FALSE;
   SEK[602].BIT.H_IN_POS1 := FALSE;
   SEK[602].BIT.H_IN_POS2 := FALSE;
   SEK[602].BIT.H_IN_POS3 := FALSE;
   SEK[602].BIT.H_IN_POS4 := FALSE;
   SEK[602].BIT.H_GR_POS := FALSE;
   SEK[602].BIT.H_SM_POS := FALSE;
   SEK[602].BIT.H_GR_POS1 := FALSE;
   SEK[602].BIT.H_SM_POS1 := FALSE;
   SEK[602].BIT.H_GR_POS2 := FALSE;
   SEK[602].BIT.H_SM_POS2 := FALSE;
   SEK[602].BIT.H_GR_POS3 := FALSE;
   SEK[602].BIT.H_SM_POS3 := FALSE;
   SEK[602].BIT.H_GR_POS4 := FALSE;
   SEK[602].BIT.H_SM_POS4 := FALSE;
   SEK[602].BIT.H_BOTTOM_POS := FALSE;
   SEK[602].BIT.H_DISABLED := FALSE;
   SEK[602].BIT.H_CLEAR := FALSE;
   SEK[602].BIT.D_MOVING_FWD := FALSE;
   SEK[602].BIT.D_MOVING_RWD := FALSE;
   SEK[602].BIT.D_RESET_AFTER := FALSE;
   SEK[602].BIT.D_PULK := FALSE;
   SEK[602].BIT.D_NO_POS := FALSE;
   SEK[602].SORTE[1] := ' ';
   SEK[602].SORTE[2] := ' ';
   SEK[602].SORTE[3] := ' ';
   SEK[602].SORTE[4] := ' ';
   SEK[602].FKT.EMS_TO_REPAIR_1 := FALSE;
   SEK[602].FKT.EMS_TO_REPAIR_2 := FALSE;
   SEK[602].FKT.EMERG_HOIST := FALSE;
   SEK[602].FKT.Reserve_03 := FALSE;
   SEK[602].FKT.EMERG_DRIVE_FC := FALSE;
   SEK[602].FKT.Reserve_05 := FALSE;
   SEK[602].FKT.LAMP_TEST := FALSE;
   SEK[602].FKT.VAC_CLEAN := FALSE;
   SEK[602].FKT.PE_TEST := FALSE;
   SEK[602].FKT.KOHLE_TEST := FALSE;
   SEK[602].FKT.KOM_TEST := FALSE;
   SEK[602].FKT.Reserve_11 := FALSE;
   SEK[602].FKT.Reserve_12 := FALSE;
   SEK[602].FKT.Reserve_13 := FALSE;
   SEK[602].FKT.Reserve_14 := FALSE;
   SEK[602].FKT.Reserve_15 := FALSE;
   SEK[602].SPARE := 16#0000;
   SEK[603].VAL.EMS_ID := 0;
   SEK[603].VAL.PROFIL := 0;
   SEK[603].VAL.DRIVE_POS := 0;
   SEK[603].VAL.HOIST_POS := 0;
   SEK[603].VAL.ERROR := 0;
   SEK[603].VAL.DRIVE_POS_PERC := 0;
   SEK[603].VAL.SEK := 0;
   SEK[603].BIT.PRESENT := FALSE;
   SEK[603].BIT.ERROR := FALSE;
   SEK[603].BIT.MAN_IR := FALSE;
   SEK[603].BIT.MORE_EMS_PRESENT := FALSE;
   SEK[603].BIT.ER_COMMAND := FALSE;
   SEK[603].BIT.W_DIST := FALSE;
   SEK[603].BIT.Spare_0_6 := FALSE;
   SEK[603].BIT.MESS_ACT := FALSE;
   SEK[603].BIT.D_MOVING := FALSE;
   SEK[603].BIT.D_NOT_MOVING := FALSE;
   SEK[603].BIT.H_MOVING := FALSE;
   SEK[603].BIT.H_NOT_MOVING := FALSE;
   SEK[603].BIT.X_MOVING := FALSE;
   SEK[603].BIT.X_NOT_MOVING := FALSE;
   SEK[603].BIT.D_IN_POS := FALSE;
   SEK[603].BIT.Spare_2_1 := FALSE;
   SEK[603].BIT.D_BEFOR_POS := FALSE;
   SEK[603].BIT.D_AFTER_POS := FALSE;
   SEK[603].BIT.D_GR_AP1 := FALSE;
   SEK[603].BIT.D_SM_AP1 := FALSE;
   SEK[603].BIT.D_GR_AP2 := FALSE;
   SEK[603].BIT.D_SM_AP2 := FALSE;
   SEK[603].BIT.H_IN_POS := FALSE;
   SEK[603].BIT.H_IN_TOPPOS := FALSE;
   SEK[603].BIT.H_IN_POS1 := FALSE;
   SEK[603].BIT.H_IN_POS2 := FALSE;
   SEK[603].BIT.H_IN_POS3 := FALSE;
   SEK[603].BIT.H_IN_POS4 := FALSE;
   SEK[603].BIT.H_GR_POS := FALSE;
   SEK[603].BIT.H_SM_POS := FALSE;
   SEK[603].BIT.H_GR_POS1 := FALSE;
   SEK[603].BIT.H_SM_POS1 := FALSE;
   SEK[603].BIT.H_GR_POS2 := FALSE;
   SEK[603].BIT.H_SM_POS2 := FALSE;
   SEK[603].BIT.H_GR_POS3 := FALSE;
   SEK[603].BIT.H_SM_POS3 := FALSE;
   SEK[603].BIT.H_GR_POS4 := FALSE;
   SEK[603].BIT.H_SM_POS4 := FALSE;
   SEK[603].BIT.H_BOTTOM_POS := FALSE;
   SEK[603].BIT.H_DISABLED := FALSE;
   SEK[603].BIT.H_CLEAR := FALSE;
   SEK[603].BIT.D_MOVING_FWD := FALSE;
   SEK[603].BIT.D_MOVING_RWD := FALSE;
   SEK[603].BIT.D_RESET_AFTER := FALSE;
   SEK[603].BIT.D_PULK := FALSE;
   // 29400 more start values not shown
END_DATA_BLOCK

DATA_BLOCK "DB_SDC_ERRORS"   // DB3722
{ S7_Optimized_Access := 'FALSE' }
AUTHOR : FFM
FAMILY : SDC
NAME : EMS_FLT
VERSION : 1.0
   VAR
      HEADER : Struct   // Struktur für Datenheader // nicht verschieben
         DB_NR : Int := 3722;   // DB Nummer
         MIN_NR_EMS : Int := 1;   // Niedrigste EMS Nummer im Daten DB
         MAX_NR_EMS : Int := 200;   // Höchste EMS Nummer im Daten DB
         START_EMS : Int := 20;   // Startadresse der EMS Daten im Daten DB
         LAENGE_EMS_StörungS : Int := 50;   // Länge Eingänge pro EMS
         ANZ_Störung_WORDS : Int := 25;   // Anzahl Störung Words
         RES12 : Int;   // Reserve
         RES14 : Int;   // Reserve
         RES16 : Int;   // Reserve
         RES18 : Int;   // Reserve
      END_STRUCT;
      EMS : Array[1..200] of Struct
         GEN_1 : Struct   // allgemeine Störung
            ER_501 : Bool;   // Störung Not Halt
            ER_502 : Bool;   // Störung Sicherung BS1FC302
            ER_503 : Bool;   // Störung EMS ID
            ER_504 : Bool;   // Störung Lebensbit
            ER_505 : Bool;   // Störung Safety-Modul KFA131 gestört (Schaltkasten)
            ER_506 : Bool;   // Reserve
            ER_507 : Bool;   // Störung Safety-Modul KFA141 gestört (Schaltkasten)
            ER_508 : Bool;   // Reserve
            ER_509 : Bool;   // Störung Profinet Fahr-FU FE1TA1
            ER_510 : Bool;   // Störung Profinet Hub-FU HE1TA1
            ER_511 : Bool;   // Störung Profinet AposOptic 1 FE1BX01
            ER_512 : Bool;   // Störung Profinet AposOptic 2 FE1BX02
            ER_513 : Bool;   // Störung Profinet Hub Seilgeber HE1GF1
            ER_514 : Bool;   // Reserve
            ER_515 : Bool;   // Störung Kommunikationsmodul BS1TFC1
            ER_516 : Bool;   // Reserve
         END_STRUCT;
         GEN_2 : Struct   // allgemeine Störung
            ER_517 : Bool;   // Störung Profinet Schwenk Drehgeber (T&R) SN1GF1
            ER_518 : Bool;   // Störung Profinet Schwenk Drehgeber (Baumer) SN1GF2
            ER_519 : Bool;   // Reserve
            ER_520 : Bool;   // Störung Profinet Schwenk-FU SN1TA1
            ER_521 : Bool;   // Reserve
            ER_522 : Bool;   // Reserve
            ER_523 : Bool;   // Reserve
            ER_524 : Bool;   // Reserve
            ER_525 : Bool;   // Störung Safety-Modul FE1TA1 gestört (Fahr-FU)
            ER_526 : Bool;   // Störung Safety-Modul HE1TA1 gestört (Hub-FU)
            ER_527 : Bool;   // Störung Safety-Modul SN1TA1 gestört (Schwenk-FU)
            ER_528 : Bool;   // Reserve
            ER_529 : Bool;   // Reserve
            ER_530 : Bool;   // Reserve
            ER_531 : Bool;   // Reserve
            ER_532 : Bool;   // Störung SPS
         END_STRUCT;
         GEN_3 : Struct   // Meldungen
            ME_801 : Bool;   // Reserve
            ME_802 : Bool;   // Reserve
            ME_803 : Bool;   // Reserve
            ME_804 : Bool;   // Reserve
            ME_805 : Bool;   // Reserve
            ME_806 : Bool;   // Reserve
            ME_807 : Bool;   // Reserve
            ME_808 : Bool;   // Reserve
            ME_809 : Bool;   // Reserve
            ME_810 : Bool;   // Reserve
            ME_811 : Bool;   // Reserve
            ME_812 : Bool;   // Reserve
            ME_813 : Bool;   // Reserve
            ME_814 : Bool;   // Reserve
            ME_815 : Bool;   // Reserve
            ME_816 : Bool;   // Reserve
         END_STRUCT;
         GEN_4 : Struct   // Meldungen
            ME_817 : Bool;   // Meldung Bypass eingeschaltet
            ME_818 : Bool;   // Meldung Initialisierung Hub
            ME_819 : Bool;   // Reserve
            ME_820 : Bool;   // Reserve
            ME_821 : Bool;   // Reserve
            ME_822 : Bool;   // Reserve
            ME_823 : Bool;   // Meldung SDC hat Betriebsart Hand angewählt
            ME_824 : Bool;   // Meldung NotAus von Anlagen-SPS
            ME_825 : Bool;   // Meldung Distanzkontrolle
            ME_826 : Bool;   // Reserve
            ME_827 : Bool;   // Reserve
            ME_828 : Bool;   // Meldung Notbetrieb ein Fahrantrieb angewählt
            ME_829 : Bool;   // Meldung Notbetrieb ein Schwenkantrieb angewählt
            ME_830 : Bool;   // Meldung Notbetrieb ohne Hub angewählt
            ME_831 : Bool;   // Meldung Notbetrieb ohne Schwenken angewählt
            ME_832 : Bool;   // Reserve
         END_STRUCT;
         DRIVE_1 : Struct   // Störungen Fahrantrieb
            ER_601 : Bool;   // Störung Fahrantrieb: Frequenzumrichter
            ER_602 : Bool;   // Reserve
            ER_603 : Bool;   // Störung Fahrantrieb: Antriebskommando nicht plausibel
            ER_604 : Bool;   // Reserve
            ER_605 : Bool;   // Reserve
            ER_606 : Bool;   // Reserve
            ER_607 : Bool;   // Störung Fahrantrieb: Geschwindigkeit zu hoch
            ER_608 : Bool;   // Störung Fahrantrieb: Geschwindigkeit zu niedrig
            ER_609 : Bool;   // Störung Fahrantrieb: Bewegung ohne Freigabe
            ER_610 : Bool;   // Störung Fahrantrieb: Positionserkennung: Sprung unzulässig
            ER_611 : Bool;   // Störung Fahrantrieb: Positionierpunkt überfahren
            ER_612 : Bool;   // Reserve
            ER_613 : Bool;   // Reserve
            ER_614 : Bool;   // Reserve
            ER_615 : Bool;   // Reserve
            ER_616 : Bool;   // Reserve
         END_STRUCT;
         DRIVE_2 : Struct   // Störungen Fahrantrieb
            ER_617 : Bool;   // Störung Fahrantrieb: APOS-Optic PN 1 status Position NIO
            ER_618 : Bool;   // Störung Fahrantrieb: APOS-Optic PN 1 status kein Positionscode erkannt
            ER_619 : Bool;   // Störung Fahrantrieb: APOS-Optic PN 1 status Position außerhalb Grenze
            ER_620 : Bool;   // Störung Fahrantrieb: APOS-Optic PN 1 status Hardware Störung
            ER_621 : Bool;   // Störung Fahrantrieb: APOS-Optic PN 1 status Temperatur Störung
            ER_622 : Bool;   // Störung Fahrantrieb: APOS-Optic PN 1 status nicht Betriebsbereit
            ER_623 : Bool;   // Störung Fahrantrieb: APOS-Optic PN 1 status Position 0
            ER_624 : Bool;   // Störung Fahrantrieb: Reserve
            ER_625 : Bool;   // Störung Fahrantrieb: APOS-Optic PN 2 status Position NIO
            ER_626 : Bool;   // Störung Fahrantrieb: APOS-Optic PN 2 status kein Positionscode erkannt
            ER_627 : Bool;   // Störung Fahrantrieb: APOS-Optic PN 2 status Position außerhalb Grenze
            ER_628 : Bool;   // Störung Fahrantrieb: APOS-Optic PN 2 status Hardware Störung
            ER_629 : Bool;   // Störung Fahrantrieb: APOS-Optic PN 2 status Temperatur Störung
            ER_630 : Bool;   // Störung Fahrantrieb: APOS-Optic PN 2 status nicht Betriebsbereit
            ER_631 : Bool;   // Störung Fahrantrieb: APOS-Optic PN 2 status Position 0
            ER_632 : Bool;   // Störung Fahrantrieb: Reserve
         END_STRUCT;
         FC_DRIVE_1 : Struct   // FU Fahrantrieb
            ER_633 : Bool;   // Störung Fahrantrieb FU 1: Überstrom
            ER_634 : Bool;   // Störung Fahrantrieb FU 1: Zwischenkreisspannung Überspannung
            ER_635 : Bool;   // Störung Fahrantrieb FU 1: Zwischenkreisspannung Unterspannung
            ER_636 : Bool;   // Störung Fahrantrieb FU 1: Übertemperatur Kühlkörper Wechselrichter
            ER_637 : Bool;   // Störung Fahrantrieb FU 1: Motordatenidentifikation fehlerhaft
            ER_638 : Bool;   // Störung Fahrantrieb FU 1: Erdschluss
            ER_639 : Bool;   // Störung Fahrantrieb FU 1: Reserve
            ER_640 : Bool;   // Störung Fahrantrieb FU 1: Führung durch PLC fehlt
            ER_641 : Bool;   // Störung Fahrantrieb FU 1: Reserve
            ER_642 : Bool;   // Störung Fahrantrieb FU 1: Reserve
            ER_643 : Bool;   // Störung Fahrantrieb FU 1: Reserve
            ER_644 : Bool;   // Störung Fahrantrieb FU 1: Reserve
            ER_645 : Bool;   // Störung Fahrantrieb FU 1: Reserve
            ER_646 : Bool;   // Störung Fahrantrieb FU 1: Reserve
            ER_647 : Bool;   // Störung Fahrantrieb FU 1: Reserve
            ER_648 : Bool;   // Störung Fahrantrieb FU 1: Reserve
         END_STRUCT;
         SAFTY_DRIVE : Struct
            ER_649 : Bool;   // Störung Fahrantrieb Safety: AposOptic 1 Sprung nicht zulässig
            ER_650 : Bool;   // Störung Fahrantrieb Safety: AposOptic 2 Sprung nicht zulässig
            ER_651 : Bool;   // Störung Fahrantrieb Safety: AposOpticwert 1 hat Limit überschritten
            ER_652 : Bool;   // Störung Fahrantrieb Safety: AposOpticwert 2 hat Limit überschritten
            ER_653 : Bool;   // Störung Fahrantrieb Safety: Geschwindigkeit AposOpticwert 1 zu hoch
            ER_654 : Bool;   // Störung Fahrantrieb Safety: Wertänderung des AposOpticwert 1 entspricht nicht der Drehrichtung
            ER_655 : Bool;   // Störung Fahrantrieb Safety: Geschwindigkeit AposOpticwert 2 zu hoch
            ER_656 : Bool;   // Störung Fahrantrieb Safety: Wertänderung des AposOpticwert 2 entspricht nicht der Drehrichtung
            ER_657 : Bool;   // Störung Fahrantrieb Safety: Not Halt Bereich nicht deffiniert
            ER_658 : Bool;   // Störung Fahrantrieb Safety: Reserve
            ER_659 : Bool;   // Störung Fahrantrieb Safety: Differenz AposOptic 1 / 2 zu hoch
            ER_660 : Bool;   // Störung Fahrantrieb Safety: Reserve
            ER_661 : Bool;   // Störung Fahrantrieb Safety: Reserve
            ER_662 : Bool;   // Störung Fahrantrieb Safety: Reserve
            ER_663 : Bool;   // Störung Fahrantrieb Safety: Reserve
            ER_664 : Bool;   // Störung Fahrantrieb Safety: Reserve
         END_STRUCT;
         FC_DRIVE_2 : Struct   // FU Fahrantrieb, Reserve
            ER_665 : Bool;   // Störung Fahrantrieb FU 2: Überstrom
            ER_666 : Bool;   // Störung Fahrantrieb FU 2: Zwischenkreisspannung Überspannung
            ER_667 : Bool;   // Störung Fahrantrieb FU 2: Zwischenkreisspannung Unterspannung
            ER_668 : Bool;   // Störung Fahrantrieb FU 2: Übertemperatur Kühlkörper Wechselrichter
            ER_669 : Bool;   // Störung Fahrantrieb FU 2: Motordatenidentifikation fehlerhaft
            ER_670 : Bool;   // Störung Fahrantrieb FU 2: Erdschluss
            ER_671 : Bool;   // Störung Fahrantrieb FU 2: Reserve
            ER_672 : Bool;   // Störung Fahrantrieb FU 2: Führung durch PLC fehlt
            ER_673 : Bool;   // Störung Fahrantrieb FU 2: Reserve
            ER_674 : Bool;   // Störung Fahrantrieb FU 2: Reserve
            ER_675 : Bool;   // Störung Fahrantrieb FU 2: Reserve
            ER_676 : Bool;   // Störung Fahrantrieb FU 2: Reserve
            ER_677 : Bool;   // Störung Fahrantrieb FU 2: Reserve
            ER_678 : Bool;   // Störung Fahrantrieb FU 2: Reserve
            ER_679 : Bool;   // Störung Fahrantrieb FU 2: Reserve
            ER_680 : Bool;   // Störung Fahrantrieb FU 2: Reserve
         END_STRUCT;
         HOIST_1 : Struct   // Störungen Hubantrieb
            ER_701 : Bool;   // Störung Hubantrieb: Frequenzumrichter
            ER_702 : Bool;   // Störung Hubantrieb: Reserve
            ER_703 : Bool;   // Störung Hubantrieb: Plausibilität Seilbruchschalter
            ER_704 : Bool;   // Störung Hubantrieb: Endlage oben erreicht
            ER_705 : Bool;   // Störung Hubantrieb: Endlage unten erreicht
            ER_706 : Bool;   // Störung Hubantrieb: Seilriss Hubseil
            ER_707 : Bool;   // Störung Hubantrieb: Reserve
            ER_708 : Bool;   // Störung Hubantrieb: Reserve
            ER_709 : Bool;   // Störung Hubantrieb: Reserve
            ER_710 : Bool;   // Störung Hubantrieb: Fangbremse und Schalter
            ER_711 : Bool;   // Störung Hubantrieb: Reserve
            ER_712 : Bool;   // Störung Hubantrieb: Reserve
            ER_713 : Bool;   // Störung Hubantrieb: Geberwert zu hoch
            ER_714 : Bool;   // Störung Hubantrieb: Geberwert zu niedrig
            ER_715 : Bool;   // Störung Hubantrieb: Hubkommando nicht plausibel
            ER_716 : Bool;   // Störung Hubantrieb: Geschwindigkeit zu hoch
         END_STRUCT;
         HOIST_2 : Struct   // Störungen Hubantrieb
            ER_717 : Bool;   // Störung Hubantrieb: Geschwindigkeit zu niedrig
            ER_718 : Bool;   // Störung Hubantrieb: Bewegung ohne Freigabe
            ER_719 : Bool;   // Störung Hubantrieb: Reserve
            ER_720 : Bool;   // Störung Hubantrieb: Sprung unzulässig
            ER_721 : Bool;   // Störung Hubantrieb: Bewegung in falsche Richtung
            ER_722 : Bool;   // Störung Hubantrieb: Referenzini nicht geschaltet
            ER_723 : Bool;   // Störung Hubantrieb: Referenzini nicht frei
            ER_724 : Bool;   // Störung Hubantrieb: Differenz Geberwerte zu groß
            ER_725 : Bool;   // Störung Hubantrieb: sichere Endlage erreicht
            ER_726 : Bool;   // Störung Hubantrieb: keine Hubfreigabe vom SDC
            ER_727 : Bool;   // Störung Hubantrieb: Reserve
            ER_728 : Bool;   // Störung Hubantrieb: Seilgeberwert fehlerhaft
            ER_729 : Bool;   // Störung Hubantrieb: G120D Positionswert fehlerhaft
            ER_730 : Bool;   // Störung Hubantrieb: Reserve
            ER_731 : Bool;   // Störung Hubantrieb: Reserve
            ER_732 : Bool;   // Störung Hubantrieb: Reserve
         END_STRUCT;
         FC_HOIST_1 : Struct   // FU Hubantrieb
            ER_733 : Bool;   // Störung Hubantrieb FU 1: Überstrom
            ER_734 : Bool;   // Störung Hubantrieb FU 1: Zwischenkreisspannung Überspannung
            ER_735 : Bool;   // Störung Hubantrieb FU 1: Zwischenkreisspannung Unterspannung
            ER_736 : Bool;   // Störung Hubantrieb FU 1: Übertemperatur Kühlkörper Wechselrichter
            ER_737 : Bool;   // Störung Hubantrieb FU 1: Motordatenidentifikation fehlerhaft
            ER_738 : Bool;   // Störung Hubantrieb FU 1: Erdschluss
            ER_739 : Bool;   // Störung Hubantrieb FU 1: Reserve
            ER_740 : Bool;   // Störung Hubantrieb FU 1: Führung durch PLC fehlt
            ER_741 : Bool;   // Störung Hubantrieb FU 1: Reserve
            ER_742 : Bool;   // Störung Hubantrieb FU 1: Reserve
            ER_743 : Bool;   // Störung Hubantrieb FU 1: Reserve
            ER_744 : Bool;   // Störung Hubantrieb FU 1: Reserve
            ER_745 : Bool;   // Störung Hubantrieb FU 1: Reserve
            ER_746 : Bool;   // Störung Hubantrieb FU 1: Reserve
            ER_747 : Bool;   // Störung Hubantrieb FU 1: Reserve
            ER_748 : Bool;   // Störung Hubantrieb FU 1: Reserve
         END_STRUCT;
         SAFTY_HOIST : Struct
            ER_749 : Bool;   // Störung Hubantrieb Safety: beide Drehrichtungen gleichzeitig angesteuert
            ER_750 : Bool;   // Störung Hubantrieb Safety: Differenz Geber 1 / 2 zu hoch
            ER_751 : Bool;   // Störung Hubantrieb Safety: Werte des Gebers 1 entsprechen nicht der Drehrichtung
            ER_752 : Bool;   // Störung Hubantrieb Safety: Werte des Gebers 2 entsprechen nicht der Drehrichtung
            ER_753 : Bool;   // Störung Hubantrieb Safety: Geschwindigkeit Geber 1 zu hoch
            ER_754 : Bool;   // Störung Hubantrieb Safety: Geschwindigkeit Geber 2 zu hoch
            ER_755 : Bool;   // Störung Hubantrieb Safety: Drehzahl des G120D entsprechen nicht der Drehrichtung
            ER_756 : Bool;   // Störung Hubantrieb Safety: Geschwindigkeit G120 Drehzahl zu hoch
            ER_757 : Bool;   // Störung Hubantrieb Safety: Positionswerte nicht gültig
            ER_758 : Bool;   // Störung Hubantrieb Safety: Referenzposition/INI nicht plausibel
            ER_759 : Bool;   // Störung Hubantrieb Safety: Durchrutschweg/Bremsweg nach Motorhaltebremse
            ER_760 : Bool;   // Störung Hubantrieb Safety: Motorhaltemoment nicht erreicht
            ER_761 : Bool;   // Störung Hubantrieb Safety: Schaltzeit Hubmagnet
            ER_762 : Bool;   // Störung Hubantrieb Safety: Plausibilität von Klinkensensoren
            ER_763 : Bool;   // Störung Hubantrieb Safety: Fangklinke hat ausgelöst
            ER_764 : Bool;   // Störung Hubantrieb Safety: Rückmeldung Safety Motor Brems Relais
         END_STRUCT;
         FC_HOIST_2 : Struct   // FU Hubantrieb, Reserve
            ER_765 : Bool;   // Störung Hubantrieb FU 2: Überstrom
            ER_766 : Bool;   // Störung Hubantrieb FU 2: Zwischenkreisspannung Überspannung
            ER_767 : Bool;   // Störung Hubantrieb FU 2: Zwischenkreisspannung Unterspannung
            ER_768 : Bool;   // Störung Hubantrieb FU 2: Übertemperatur Kühlkörper Wechselrichter
            ER_769 : Bool;   // Störung Hubantrieb FU 2: Motordatenidentifikation fehlerhaft
            ER_770 : Bool;   // Störung Hubantrieb FU 2: Erdschluss
            ER_771 : Bool;   // Störung Hubantrieb FU 2: Reserve
            ER_772 : Bool;   // Störung Hubantrieb FU 2: Führung durch PLC fehlt
            ER_773 : Bool;   // Störung Hubantrieb FU 2: Reserve
            ER_774 : Bool;   // Störung Hubantrieb FU 2: Reserve
            ER_775 : Bool;   // Störung Hubantrieb FU 2: Reserve
            ER_776_ : Bool;   // Störung Hubantrieb FU 2: Reserve
            ER_777 : Bool;   // Störung Hubantrieb FU 2: Reserve
            ER_778 : Bool;   // Störung Hubantrieb FU 2: Reserve
            ER_779 : Bool;   // Störung Hubantrieb FU 2: Reserve
            ER_780 : Bool;   // Störung Hubantrieb FU 2: Reserve
         END_STRUCT;
         Reserve_1 : Struct
            ER_401 : Bool;   // Reserve
            ER_402 : Bool;   // Reserve
            ER_403 : Bool;   // Reserve
            ER_404 : Bool;   // Reserve
            ER_405 : Bool;   // Reserve
            ER_406 : Bool;   // Reserve
            ER_407 : Bool;   // Reserve
            ER_408 : Bool;   // Reserve
            ER_409 : Bool;   // Reserve
            ER_410 : Bool;   // Reserve
            ER_411 : Bool;   // Reserve
            ER_412 : Bool;   // Reserve
            ER_413 : Bool;   // Reserve
            ER_414 : Bool;   // Reserve
            ER_415 : Bool;   // Reserve
            ER_416 : Bool;   // Reserve
         END_STRUCT;
         Reserve_2 : Struct
            ER_417 : Bool;   // Reserve
            ER_418 : Bool;   // Reserve
            ER_419 : Bool;   // Reserve
            ER_420 : Bool;   // Reserve
            ER_421 : Bool;   // Reserve
            ER_422 : Bool;   // Reserve
            ER_423 : Bool;   // Reserve
            ER_424 : Bool;   // Reserve
            ER_425 : Bool;   // Reserve
            ER_426 : Bool;   // Reserve
            ER_427 : Bool;   // Reserve
            ER_428 : Bool;   // Reserve
            ER_429 : Bool;   // Reserve
            ER_430 : Bool;   // Reserve
            ER_431 : Bool;   // Reserve
            ER_432 : Bool;   // Reserve
         END_STRUCT;
         Reserve_3 : Struct
            ER_433 : Bool;   // Reserve
            ER_434 : Bool;   // Reserve
            ER_435 : Bool;   // Reserve
            ER_436 : Bool;   // Reserve
            ER_437 : Bool;   // Reserve
            ER_438 : Bool;   // Reserve
            ER_439 : Bool;   // Reserve
            ER_440 : Bool;   // Reserve
            ER_441 : Bool;   // Reserve
            ER_442 : Bool;   // Reserve
            ER_443 : Bool;   // Reserve
            ER_444 : Bool;   // Reserve
            ER_445 : Bool;   // Reserve
            ER_446 : Bool;   // Reserve
            ER_447 : Bool;   // Reserve
            ER_448 : Bool;   // Reserve
         END_STRUCT;
         Reserve_4 : Struct
            ER_449 : Bool;   // Reserve
            ER_450 : Bool;   // Reserve
            ER_451 : Bool;   // Reserve
            ER_452 : Bool;   // Reserve
            ER_453 : Bool;   // Reserve
            ER_454 : Bool;   // Reserve
            ER_455 : Bool;   // Reserve
            ER_456 : Bool;   // Reserve
            ER_457 : Bool;   // Reserve
            ER_458 : Bool;   // Reserve
            ER_459 : Bool;   // Reserve
            ER_460 : Bool;   // Reserve
            ER_461 : Bool;   // Reserve
            ER_462 : Bool;   // Reserve
            ER_463 : Bool;   // Reserve
            ER_464 : Bool;   // Reserve